(* Logix 5000 project; controller OWF Emulate 5570 rev 30.12; software revision 30.00; part 2 of 4 *)
(* tags used below, declared in another part *)
   OWF_Key : DINT[512,17];
   OWF_Ver : DINT;
(* MainProgram, continued *)

   	OWF_Key[185,11]:=700678053;
   	OWF_Key[185,12]:=1316216993;
   	OWF_Key[186,9]:=1263200427;
   	OWF_Key[186,10]:=1232581124;
   	OWF_Key[186,11]:=662303121;
   	OWF_Key[186,12]:=704428579;
   	OWF_Key[187,9]:=902189893;
   	OWF_Key[187,10]:=650291179;
   	OWF_Key[187,11]:=622514985;
   	OWF_Key[187,12]:=885208114;
   	OWF_Key[188,9]:=1740254790;
   	OWF_Key[188,10]:=19492587;
   	OWF_Key[188,11]:=1358355453;
   	OWF_Key[188,12]:=43227168;
   	OWF_Key[189,9]:=341427661;
   	OWF_Key[189,10]:=237281733;
   	OWF_Key[189,11]:=1752374772;
   	OWF_Key[189,12]:=1623944067;
   	OWF_Key[190,9]:=1165233075;
   	OWF_Key[190,10]:=2098490866;
   	OWF_Key[190,11]:=1663872531;
   	OWF_Key[190,12]:=1678946563;
   	OWF_Key[191,9]:=828491605;
   	OWF_Key[191,10]:=1917075649;
   	OWF_Key[191,11]:=1124953821;
   	OWF_Key[191,12]:=1041503626;
   	OWF_Key[192,9]:=1689318782;
   	OWF_Key[192,10]:=1423675752;
   	OWF_Key[192,11]:=512282933;
   	OWF_Key[192,12]:=918312780;
   	OWF_Key[193,9]:=417565917;
   	OWF_Key[193,10]:=588616254;
   	OWF_Key[193,11]:=933238473;
   	OWF_Key[193,12]:=1518544589;
   	OWF_Key[194,9]:=511552150;
   	OWF_Key[194,10]:=1772464712;
   	OWF_Key[194,11]:=1163529062;
   	OWF_Key[194,12]:=675427433;
   	OWF_Key[195,9]:=886772734;
   	OWF_Key[195,10]:=872507846;
   	OWF_Key[195,11]:=1433255703;
   	OWF_Key[195,12]:=78408779;
   	OWF_Key[196,9]:=1967144636;
   	OWF_Key[196,10]:=2114794010;
   	OWF_Key[196,11]:=937696784;
   	OWF_Key[196,12]:=1841817725;
   	OWF_Key[197,9]:=543733851;
   	OWF_Key[197,10]:=1472607323;
   	OWF_Key[197,11]:=1881437884;
   	OWF_Key[197,12]:=1635644016;
   	OWF_Key[198,9]:=606394668;
   	OWF_Key[198,10]:=379369195;
   	OWF_Key[198,11]:=1444811109;
   	OWF_Key[198,12]:=1865415747;
   	OWF_Key[199,9]:=73384272;
   	OWF_Key[199,10]:=318304038;
   	OWF_Key[199,11]:=1072391895;
   	OWF_Key[199,12]:=257743095;
   	OWF_Key[200,9]:=1376967215;
   	OWF_Key[200,10]:=286485900;
   	OWF_Key[200,11]:=1302123460;
   	OWF_Key[200,12]:=1695542832;
   	OWF_Key[201,9]:=1565873958;
   	OWF_Key[201,10]:=1658681123;
   	OWF_Key[201,11]:=869814778;
   	OWF_Key[201,12]:=1614127583;
   	OWF_Key[202,9]:=1442184069;
   	OWF_Key[202,10]:=1378673233;
   	OWF_Key[202,11]:=367634315;
   	OWF_Key[202,12]:=749842782;
   	OWF_Key[203,9]:=358016958;
   	OWF_Key[203,10]:=1331305300;
   	OWF_Key[203,11]:=1285755694;
   	OWF_Key[203,12]:=1076068166;
   	OWF_Key[204,9]:=708598934;
   	OWF_Key[204,10]:=2016392191;
   	OWF_Key[204,11]:=54308888;
   	OWF_Key[204,12]:=1057259517;
   	OWF_Key[205,9]:=203186814;
   	OWF_Key[205,10]:=794532971;
   	OWF_Key[205,11]:=1428669067;
   	OWF_Key[205,12]:=1461313202;
   	OWF_Key[206,9]:=1784635668;
   	OWF_Key[206,10]:=710140484;
   	OWF_Key[206,11]:=67224826;
   	OWF_Key[206,12]:=437768377;
   	OWF_Key[207,9]:=2035750048;
   	OWF_Key[207,10]:=384041580;
   	OWF_Key[207,11]:=296753188;
   	OWF_Key[207,12]:=1785547776;
   	OWF_Key[208,9]:=1478080033;
   	OWF_Key[208,10]:=2029658272;
   	OWF_Key[208,11]:=707257918;
   	OWF_Key[208,12]:=1299161440;
   	OWF_Key[209,9]:=1393054311;
   	OWF_Key[209,10]:=1894932492;
   	OWF_Key[209,11]:=619202765;
   	OWF_Key[209,12]:=189108264;
   	OWF_Key[210,9]:=1572386515;
   	OWF_Key[210,10]:=1828673857;
   	OWF_Key[210,11]:=1993473823;
   	OWF_Key[210,12]:=73594153;
   	OWF_Key[211,9]:=1184769439;
   	OWF_Key[211,10]:=1936440244;
   	OWF_Key[211,11]:=935061554;
   	OWF_Key[211,12]:=149096850;
   	OWF_Key[212,9]:=1900216788;
   	OWF_Key[212,10]:=56648648;
   	OWF_Key[212,11]:=1184648305;
   	OWF_Key[212,12]:=778107636;
   	OWF_Key[213,9]:=263723127;
   	OWF_Key[213,10]:=1061340316;
   	OWF_Key[213,11]:=1706699901;
   	OWF_Key[213,12]:=851139445;
   	OWF_Key[214,9]:=1866191994;
   	OWF_Key[214,10]:=1265826094;
   	OWF_Key[214,11]:=1893173788;
   	OWF_Key[214,12]:=1185508622;
   	OWF_Key[215,9]:=432963339;
   	OWF_Key[215,10]:=930912264;
   	OWF_Key[215,11]:=1473487116;
   	OWF_Key[215,12]:=1240528203;
   	OWF_Key[216,9]:=832362750;
   	OWF_Key[216,10]:=53435343;
   	OWF_Key[216,11]:=473043438;
   	OWF_Key[216,12]:=76142584;
   	OWF_Key[217,9]:=866996792;
   	OWF_Key[217,10]:=825249854;
   	OWF_Key[217,11]:=986453816;
   	OWF_Key[217,12]:=1455610264;
   	OWF_Key[218,9]:=1923606857;
   	OWF_Key[218,10]:=1160389397;
   	OWF_Key[218,11]:=167392645;
   	OWF_Key[218,12]:=761527794;
   	OWF_Key[219,9]:=1345872227;
   	OWF_Key[219,10]:=1835824993;
   	OWF_Key[219,11]:=1850219615;
   	OWF_Key[219,12]:=2124120876;
   	OWF_Key[220,9]:=605851105;
   	OWF_Key[220,10]:=962199035;
   	OWF_Key[220,11]:=706661987;
   	OWF_Key[220,12]:=157680519;
   	OWF_Key[221,9]:=1484271236;
   	OWF_Key[221,10]:=562747976;
   	OWF_Key[221,11]:=1031426104;
   	OWF_Key[221,12]:=2014277938;
   	OWF_Key[222,9]:=1518806301;
   	OWF_Key[222,10]:=1196972058;
   	OWF_Key[222,11]:=834756739;
   	OWF_Key[222,12]:=1825620384;
   	OWF_Key[223,9]:=1107633867;
   	OWF_Key[223,10]:=844435349;
   	OWF_Key[223,11]:=101438149;
   	OWF_Key[223,12]:=274480237;
   	OWF_Key[224,9]:=330594083;
   	OWF_Key[224,10]:=851981438;
   	OWF_Key[224,11]:=734730016;
   	OWF_Key[224,12]:=1622996730;
   	OWF_Key[225,9]:=509439923;
   	OWF_Key[225,10]:=488128788;
   	OWF_Key[225,11]:=321219229;
   	OWF_Key[225,12]:=115663854;
   	OWF_Key[226,9]:=319922320;
   	OWF_Key[226,10]:=32596412;
   	OWF_Key[226,11]:=600946799;
   	OWF_Key[226,12]:=789183496;
   	OWF_Key[227,9]:=1575599257;
   	OWF_Key[227,10]:=509704494;
   	OWF_Key[227,11]:=320400967;
   	OWF_Key[227,12]:=90882807;
   	OWF_Key[228,9]:=67010183;
   	OWF_Key[228,10]:=1430271682;
   	OWF_Key[228,11]:=1541114392;
   	OWF_Key[228,12]:=486872836;
   	OWF_Key[229,9]:=1985386453;
   	OWF_Key[229,10]:=743916993;
   	OWF_Key[229,11]:=1038816091;
   	OWF_Key[229,12]:=1128633452;
   	OWF_Key[230,9]:=1230507347;
   	OWF_Key[230,10]:=204341659;
   	OWF_Key[230,11]:=1327761903;
   	OWF_Key[230,12]:=1110131463;
   	OWF_Key[231,9]:=875175521;
   	OWF_Key[231,10]:=831829301;
   	OWF_Key[231,11]:=729903640;
   	OWF_Key[231,12]:=1342317219;
   	OWF_Key[232,9]:=735217235;
   	OWF_Key[232,10]:=25404189;
   	OWF_Key[232,11]:=1924349757;
   	OWF_Key[232,12]:=1726880295;
   	OWF_Key[233,9]:=617710046;
   	OWF_Key[233,10]:=1997859713;
   	OWF_Key[233,11]:=1355438325;
   	OWF_Key[233,12]:=1453957869;
   	OWF_Key[234,9]:=370548099;
   	OWF_Key[234,10]:=452260747;
   	OWF_Key[234,11]:=954206997;
   	OWF_Key[234,12]:=1617031508;
   	OWF_Key[235,9]:=220384771;
   	OWF_Key[235,10]:=369121378;
   	OWF_Key[235,11]:=1735385215;
   	OWF_Key[235,12]:=1555781138;
   	OWF_Key[236,9]:=975725139;
   	OWF_Key[236,10]:=1267496554;
   	OWF_Key[236,11]:=1256808528;
   	OWF_Key[236,12]:=1819055267;
   	OWF_Key[237,9]:=732173551;
   	OWF_Key[237,10]:=513189099;
   	OWF_Key[237,11]:=1913299098;
   	OWF_Key[237,12]:=1166272901;
   	OWF_Key[238,9]:=976841642;
   	OWF_Key[238,10]:=1662757885;
   	OWF_Key[238,11]:=788281835;
   	OWF_Key[238,12]:=348319935;
   	OWF_Key[239,9]:=1485357753;
   	OWF_Key[239,10]:=2125315212;
   	OWF_Key[239,11]:=712191996;
   	OWF_Key[239,12]:=1015872871;
   	OWF_Key[240,9]:=636618036;
   	OWF_Key[240,10]:=1156635726;
   	OWF_Key[240,11]:=312419555;
   	OWF_Key[240,12]:=1171231843;
   	OWF_Key[241,9]:=760182292;
   	OWF_Key[241,10]:=1638351670;
   	OWF_Key[241,11]:=1089247529;
   	OWF_Key[241,12]:=92018885;
   	OWF_Key[242,9]:=951060119;
   	OWF_Key[242,10]:=587755415;
   	OWF_Key[242,11]:=1572914183;
   	OWF_Key[242,12]:=530552876;
   	OWF_Key[243,9]:=1521645385;
   	OWF_Key[243,10]:=563714124;
   	OWF_Key[243,11]:=1320117927;
   	OWF_Key[243,12]:=499630181;
   	OWF_Key[244,9]:=443279081;
   	OWF_Key[244,10]:=459094614;
   	OWF_Key[244,11]:=429852943;
   	OWF_Key[244,12]:=1357255337;
   	OWF_Key[245,9]:=2126590490;
   	OWF_Key[245,10]:=958701753;
   	OWF_Key[245,11]:=1694545154;
   	OWF_Key[245,12]:=1699505041;
   	OWF_Key[246,9]:=714967445;
   	OWF_Key[246,10]:=818909417;
   	OWF_Key[246,11]:=2000705415;
   	OWF_Key[246,12]:=812175043;
   	OWF_Key[247,9]:=690539805;
   	OWF_Key[247,10]:=320296430;
   	OWF_Key[247,11]:=2088794569;
   	OWF_Key[247,12]:=2048851186;
   	OWF_Key[248,9]:=1418362003;
   	OWF_Key[248,10]:=772738491;
   	OWF_Key[248,11]:=608671834;
   	OWF_Key[248,12]:=1563232568;
   	OWF_Key[249,9]:=1992968931;
   	OWF_Key[249,10]:=443260534;
   	OWF_Key[249,11]:=475757846;
   	OWF_Key[249,12]:=690073579;
   	OWF_Key[250,9]:=1125311706;
   	OWF_Key[250,10]:=1050444347;
   	OWF_Key[250,11]:=77048878;
   	OWF_Key[250,12]:=1221726213;
   	OWF_Key[251,9]:=23263864;
   	OWF_Key[251,10]:=817695650;
   	OWF_Key[251,11]:=238910220;
   	OWF_Key[251,12]:=1101491130;
   	OWF_Key[252,9]:=849558070;
   	OWF_Key[252,10]:=1729978099;
   	OWF_Key[252,11]:=351451070;
   	OWF_Key[252,12]:=1932474899;
   	OWF_Key[253,9]:=1716607782;
   	OWF_Key[253,10]:=597806638;
   	OWF_Key[253,11]:=594517253;
   	OWF_Key[253,12]:=1313352884;
   	OWF_Key[254,9]:=1389320638;
   	OWF_Key[254,10]:=1479710077;
   	OWF_Key[254,11]:=39152000;
   	OWF_Key[254,12]:=1262503749;
   	OWF_Key[255,9]:=523479812;
   	OWF_Key[255,10]:=730328114;
   	OWF_Key[255,11]:=1256933613;
   	OWF_Key[255,12]:=832190698;
   	OWF_Key[256,0]:=1909298189;
   	OWF_Key[256,1]:=179491594;
   	OWF_Key[256,2]:=930979855;
   	OWF_Key[256,3]:=1826970333;
   	OWF_Key[256,4]:=2108067730;
   	OWF_Key[256,5]:=1321930337;
   	OWF_Key[256,6]:=1292378578;
   	OWF_Key[256,7]:=528139296;
   	OWF_Key[256,8]:=1454317303;
   	OWF_Key[256,9]:=1411726950;
   	OWF_Key[256,10]:=760872820;
   	OWF_Key[256,11]:=1454011296;
   	OWF_Key[256,12]:=1435946443;
   	OWF_Key[257,0]:=2080112384;
   	OWF_Key[257,1]:=2058516218;
   	OWF_Key[257,2]:=201781603;
   	OWF_Key[257,3]:=974822888;
   	OWF_Key[257,4]:=913739450;
   	OWF_Key[257,5]:=255145122;
   	OWF_Key[257,6]:=1164040444;
   	OWF_Key[257,7]:=1649300770;
   	OWF_Key[257,8]:=1308958305;
   	OWF_Key[257,9]:=1833316665;
   	OWF_Key[257,10]:=965533626;
   	OWF_Key[257,11]:=1955596663;
   	OWF_Key[257,12]:=756111181;
   	OWF_Key[258,0]:=188290248;
   	OWF_Key[258,1]:=1487618761;
   	OWF_Key[258,2]:=1152942549;
   	OWF_Key[258,3]:=647319114;
   	OWF_Key[258,4]:=1246205489;
   	OWF_Key[258,5]:=190536859;
   	OWF_Key[258,6]:=1474452229;
   	OWF_Key[258,7]:=1211715374;
   	OWF_Key[258,8]:=996148662;
   	OWF_Key[258,9]:=40987582;
   	OWF_Key[258,10]:=2113307878;
   	OWF_Key[258,11]:=79456365;
   	OWF_Key[258,12]:=1496771068;
   	OWF_Key[259,0]:=1771169746;
   	OWF_Key[259,1]:=1499571985;
   	OWF_Key[259,2]:=182288128;
   	OWF_Key[259,3]:=787798492;
   	OWF_Key[259,4]:=2049043781;
   	OWF_Key[259,5]:=971867535;
   	OWF_Key[259,6]:=353694007;
   	OWF_Key[259,7]:=1196884289;
   	OWF_Key[259,8]:=469754060;
   	OWF_Key[259,9]:=1351904685;
   	OWF_Key[259,10]:=776834163;
   	OWF_Key[259,11]:=563849352;
   	OWF_Key[259,12]:=1687317924;
   	OWF_Key[260,0]:=197268257;
   	OWF_Key[260,1]:=1562397221;
   	OWF_Key[260,2]:=1268651049;
   	OWF_Key[260,3]:=2000952175;
   	OWF_Key[260,4]:=1561123196;
   	OWF_Key[260,5]:=1239508018;
   	OWF_Key[260,6]:=1278308208;
   	OWF_Key[260,7]:=2137033599;
   	OWF_Key[260,8]:=706681873;
   	OWF_Key[260,9]:=1531967027;
   	OWF_Key[260,10]:=1582992287;
   	OWF_Key[260,11]:=1589667041;
   	OWF_Key[260,12]:=1632710709;
   	OWF_Key[261,0]:=1713243906;
   	OWF_Key[261,1]:=456764431;
   	OWF_Key[261,2]:=1285431790;
   	OWF_Key[261,3]:=1056490938;
   	OWF_Key[261,4]:=443278195;
   	OWF_Key[261,5]:=655715940;
   	OWF_Key[261,6]:=474288957;
   	OWF_Key[261,7]:=743704672;
   	OWF_Key[261,8]:=1032636258;
   	OWF_Key[261,9]:=1982657051;
   	OWF_Key[261,10]:=1461505893;
   	OWF_Key[261,11]:=1251097594;
   	OWF_Key[261,12]:=1893699385;
   	OWF_Key[262,0]:=727961623;
   	OWF_Key[262,1]:=479034231;
   	OWF_Key[262,2]:=1801422076;
   	OWF_Key[262,3]:=97476380;
   	OWF_Key[262,4]:=1502493348;
   	OWF_Key[262,5]:=925680604;
   	OWF_Key[262,6]:=1129443202;
   	OWF_Key[262,7]:=1551038546;
   	OWF_Key[262,8]:=2014591270;
   	OWF_Key[262,9]:=1190072555;
   	OWF_Key[262,10]:=742299502;
   	OWF_Key[262,11]:=152374670;
   	OWF_Key[262,12]:=1358004664;
   	OWF_Key[263,0]:=1665333302;
   	OWF_Key[263,1]:=1728497092;
   	OWF_Key[263,2]:=1506278205;
   	OWF_Key[263,3]:=1554919913;
   	OWF_Key[263,4]:=654676244;
   	OWF_Key[263,5]:=938138664;
   	OWF_Key[263,6]:=1695588185;
   	OWF_Key[263,7]:=1018196095;
   	OWF_Key[263,8]:=926711657;
   	OWF_Key[263,9]:=1698779979;
   	OWF_Key[263,10]:=1903955519;
   	OWF_Key[263,11]:=656400961;
   	OWF_Key[263,12]:=1092404117;
   	OWF_Key[264,0]:=1265871845;
   	OWF_Key[264,1]:=1310650858;
   	OWF_Key[264,2]:=1110441492;
   	OWF_Key[264,3]:=64254185;
   	OWF_Key[264,4]:=71092357;
   	OWF_Key[264,5]:=911339644;
   	OWF_Key[264,6]:=910281411;
   	OWF_Key[264,7]:=701064343;
   	OWF_Key[264,8]:=280054373;
   	OWF_Key[264,9]:=1999806079;
   	OWF_Key[264,10]:=1856194407;
   	OWF_Key[264,11]:=2106992576;
   	OWF_Key[264,12]:=1848449120;
   	OWF_Key[265,0]:=1444563459;
   	OWF_Key[265,1]:=377741508;
   	OWF_Key[265,2]:=424778512;
   	OWF_Key[265,3]:=847388549;
   	OWF_Key[265,4]:=210722876;
   	OWF_Key[265,5]:=244777580;
   	OWF_Key[265,6]:=1835771034;
   	OWF_Key[265,7]:=520328668;
   	OWF_Key[265,8]:=1590554406;
   	OWF_Key[265,9]:=2014826841;
   	OWF_Key[265,10]:=984893395;
   	OWF_Key[265,11]:=1242446533;
   	OWF_Key[265,12]:=729667471;
   	OWF_Key[266,0]:=1330920216;
   	OWF_Key[266,1]:=2073347181;
   	OWF_Key[266,2]:=623283799;
   	OWF_Key[266,3]:=668461211;
   	OWF_Key[266,4]:=2068984788;
   	OWF_Key[266,5]:=1869166776;
   	OWF_Key[266,6]:=1675179723;
   	OWF_Key[266,7]:=171657924;
   	OWF_Key[266,8]:=2006816936;
   	OWF_Key[266,9]:=1771515439;
   	OWF_Key[266,10]:=1458869826;
   	OWF_Key[266,11]:=2126885731;
   	OWF_Key[266,12]:=446766808;
   	OWF_Key[267,0]:=723153773;
   	OWF_Key[267,1]:=1434115044;
   	OWF_Key[267,2]:=982028123;
   	OWF_Key[267,3]:=2017097021;
   	OWF_Key[267,4]:=928613763;
   	OWF_Key[267,5]:=1267329486;
   	OWF_Key[267,6]:=888233137;
   	OWF_Key[267,7]:=323445376;
   	OWF_Key[267,8]:=2120266118;
   	OWF_Key[267,9]:=699690438;
   	OWF_Key[267,10]:=1851502649;
   	OWF_Key[267,11]:=1879659818;
   	OWF_Key[267,12]:=63749953;
   	OWF_Key[268,0]:=1191293725;
   	OWF_Key[268,1]:=1242872285;
   	OWF_Key[268,2]:=1704548290;
   	OWF_Key[268,3]:=131127079;
   	OWF_Key[268,4]:=112917177;
   	OWF_Key[268,5]:=2082559947;
   	OWF_Key[268,6]:=1804396835;
   	OWF_Key[268,7]:=1736270177;
   	OWF_Key[268,8]:=1447868554;
   	OWF_Key[268,9]:=116578103;
   	OWF_Key[268,10]:=123670109;
   	OWF_Key[268,11]:=225035136;
   	OWF_Key[268,12]:=494051068;
   	OWF_Key[269,0]:=981365361;
   	OWF_Key[269,1]:=356297074;
   	OWF_Key[269,2]:=1178165977;
   	OWF_Key[269,3]:=925717798;
   	OWF_Key[269,4]:=1579250891;
   	OWF_Key[269,5]:=1909207467;
   	OWF_Key[269,6]:=364488170;
   	OWF_Key[269,7]:=1991543628;
   	OWF_Key[269,8]:=539128452;
   	OWF_Key[269,9]:=1418683480;
   	OWF_Key[269,10]:=1741862447;
   	OWF_Key[269,11]:=288771385;
   	OWF_Key[269,12]:=2100436399;
   	OWF_Key[270,0]:=807771279;
   	OWF_Key[270,1]:=38360465;
   	OWF_Key[270,2]:=325622113;
   	OWF_Key[270,3]:=384307439;
   	OWF_Key[270,4]:=935251297;
   	OWF_Key[270,5]:=1358532483;
   	OWF_Key[270,6]:=1161114543;
   	OWF_Key[270,7]:=897783333;
   	OWF_Key[270,8]:=1210966455;
   	OWF_Key[270,9]:=690422852;
   	OWF_Key[270,10]:=1210663776;
   	OWF_Key[270,11]:=1615774481;
   	OWF_Key[270,12]:=121890596;
   	OWF_Key[271,0]:=420087205;
   	OWF_Key[271,1]:=6570589;
   	OWF_Key[271,2]:=1677029070;
   	OWF_Key[271,3]:=1171283268;
   	OWF_Key[271,4]:=151669090;
   	OWF_Key[271,5]:=1610835874;
   	OWF_Key[271,6]:=1049960611;
   	OWF_Key[271,7]:=1011567790;
   	OWF_Key[271,8]:=1506255067;
   	OWF_Key[271,9]:=88410857;
   	OWF_Key[271,10]:=566557477;
   	OWF_Key[271,11]:=577114258;
   	OWF_Key[271,12]:=507847073;
   	OWF_Key[272,0]:=1130841498;
   	OWF_Key[272,1]:=1208532936;
   	OWF_Key[272,2]:=2083516122;
   	OWF_Key[272,3]:=997587375;
   	OWF_Key[272,4]:=446553888;
   	OWF_Key[272,5]:=1458442193;
   	OWF_Key[272,6]:=2097366676;
   	OWF_Key[272,7]:=365072649;
   	OWF_Key[272,8]:=609768654;
   	OWF_Key[272,9]:=1628492900;
   	OWF_Key[272,10]:=661311241;
   	OWF_Key[272,11]:=2061825909;
   	OWF_Key[272,12]:=982939224;
   	OWF_Key[273,0]:=1432208058;
   	OWF_Key[273,1]:=1611062291;
   	OWF_Key[273,2]:=53505219;
   	OWF_Key[273,3]:=1410831432;
   	OWF_Key[273,4]:=1603737596;
   	OWF_Key[273,5]:=2006606228;
   	OWF_Key[273,6]:=1702403367;
   	OWF_Key[273,7]:=2024779983;
   	OWF_Key[273,8]:=1642019509;
   	OWF_Key[273,9]:=1410195440;
   	OWF_Key[273,10]:=619437922;
   	OWF_Key[273,11]:=1211109155;
   	OWF_Key[273,12]:=866002016;
   	OWF_Key[274,0]:=581115914;
   	OWF_Key[274,1]:=1418969672;
   	OWF_Key[274,2]:=2060980742;
   	OWF_Key[274,3]:=754371406;
   	OWF_Key[274,4]:=608644476;
   	OWF_Key[274,5]:=759310711;
   	OWF_Key[274,6]:=777736275;
   	OWF_Key[274,7]:=1865828594;
   	OWF_Key[274,8]:=1641635049;
   	OWF_Key[274,9]:=41710555;
   	OWF_Key[274,10]:=755866891;
   	OWF_Key[274,11]:=1067621783;
   	OWF_Key[274,12]:=85169824;
   	OWF_Key[275,0]:=1852880267;
   	OWF_Key[275,1]:=973223475;
   	OWF_Key[275,2]:=1020637725;
   	OWF_Key[275,3]:=2132448151;
   	OWF_Key[275,4]:=1863827790;
   	OWF_Key[275,5]:=1183600567;
   	OWF_Key[275,6]:=355277438;
   	OWF_Key[275,7]:=1331619337;
   	OWF_Key[275,8]:=320631388;
   	OWF_Key[275,9]:=743910291;
   	OWF_Key[275,10]:=1485471229;
   	OWF_Key[275,11]:=2052565943;
   	OWF_Key[275,12]:=134289450;
   	OWF_Key[276,0]:=1358205830;
   	OWF_Key[276,1]:=94720866;
   	OWF_Key[276,2]:=1006129356;
   	OWF_Key[276,3]:=45328915;
   	OWF_Key[276,4]:=2063960286;
   	OWF_Key[276,5]:=1824801631;
   	OWF_Key[276,6]:=1997963052;
   	OWF_Key[276,7]:=1976531471;
   	OWF_Key[276,8]:=1047041442;
   	OWF_Key[276,9]:=1147595151;
   	OWF_Key[276,10]:=1532494885;
   	OWF_Key[276,11]:=541152753;
   	OWF_Key[276,12]:=1911908976;
   	OWF_Key[277,0]:=1376252338;
   	OWF_Key[277,1]:=269498259;
   	OWF_Key[277,2]:=1522115671;
   	OWF_Key[277,3]:=152049218;
   	OWF_Key[277,4]:=1299952226;
   	OWF_Key[277,5]:=1699600321;
   	OWF_Key[277,6]:=1198368614;
   	OWF_Key[277,7]:=1031693347;
   	OWF_Key[277,8]:=566771635;
   	OWF_Key[277,9]:=759840169;
   	OWF_Key[277,10]:=530325796;
   	OWF_Key[277,11]:=103291625;
   	OWF_Key[277,12]:=885409307;
   	OWF_Key[278,0]:=1328624873;
   	OWF_Key[278,1]:=1823532889;
   	OWF_Key[278,2]:=2086426509;
   	OWF_Key[278,3]:=1050375054;
   	OWF_Key[278,4]:=680213368;
   	OWF_Key[278,5]:=1611291071;
   	OWF_Key[278,6]:=1233222043;
   	OWF_Key[278,7]:=978756704;
   	OWF_Key[278,8]:=218500436;
   	OWF_Key[278,9]:=1064704980;
   	OWF_Key[278,10]:=2018975882;
   	OWF_Key[278,11]:=1792732229;
   	OWF_Key[278,12]:=1925215460;
   	OWF_Key[279,0]:=1715027586;
   	OWF_Key[279,1]:=935390411;
   	OWF_Key[279,2]:=1409344007;
   	OWF_Key[279,3]:=736299114;
   	OWF_Key[279,4]:=473416930;
   	OWF_Key[279,5]:=573329454;
   	OWF_Key[279,6]:=299400874;
   	OWF_Key[279,7]:=780542717;
   	OWF_Key[279,8]:=1932949313;
   	OWF_Key[279,9]:=1152271737;
   	OWF_Key[279,10]:=1913736579;
   	OWF_Key[279,11]:=439032107;
   	OWF_Key[279,12]:=2064816898;
   	OWF_Key[280,0]:=570567511;
   	OWF_Key[280,1]:=1114156889;
   	OWF_Key[280,2]:=709066882;
   	OWF_Key[280,3]:=878708860;
   	OWF_Key[280,4]:=1852019797;
   	OWF_Key[280,5]:=54158267;
   	OWF_Key[280,6]:=1712298224;
   	OWF_Key[280,7]:=672377733;
   	OWF_Key[280,8]:=795609163;
   	OWF_Key[280,9]:=1138980779;
   	OWF_Key[280,10]:=601731358;
   	OWF_Key[280,11]:=1532096588;
   	OWF_Key[280,12]:=1333532316;
   	OWF_Key[281,0]:=2398887;
   	OWF_Key[281,1]:=2103211707;
   	OWF_Key[281,2]:=1187423234;
   	OWF_Key[281,3]:=2115109801;
   	OWF_Key[281,4]:=204920429;
   	OWF_Key[281,5]:=777528471;
   	OWF_Key[281,6]:=44267019;
   	OWF_Key[281,7]:=1009268664;
   	OWF_Key[281,8]:=760040378;
   	OWF_Key[281,9]:=696947813;
   	OWF_Key[281,10]:=1708996504;
   	OWF_Key[281,11]:=1107831299;
   	OWF_Key[281,12]:=838778621;
   	OWF_Key[282,0]:=2094710692;
   	OWF_Key[282,1]:=199333410;
   	OWF_Key[282,2]:=143625877;
   	OWF_Key[282,3]:=742121388;
   	OWF_Key[282,4]:=395971221;
   	OWF_Key[282,5]:=498064101;
   	OWF_Key[282,6]:=592008830;
   	OWF_Key[282,7]:=1676658099;
   	OWF_Key[282,8]:=2073316084;
   	OWF_Key[282,9]:=775722435;
   	OWF_Key[282,10]:=1942183518;
   	OWF_Key[282,11]:=493527397;
   	OWF_Key[282,12]:=480575079;
   	OWF_Key[283,0]:=455375500;
   	OWF_Key[283,1]:=128497964;
   	OWF_Key[283,2]:=1573282074;
   	OWF_Key[283,3]:=59351966;
   	OWF_Key[283,4]:=274174963;
   	OWF_Key[283,5]:=148866559;
   	OWF_Key[283,6]:=1070692901;
   	OWF_Key[283,7]:=1149677535;
   	OWF_Key[283,8]:=643615893;
   	OWF_Key[283,9]:=458736794;
   	OWF_Key[283,10]:=1074207849;
   	OWF_Key[283,11]:=1880670902;
   	OWF_Key[283,12]:=954610762;
   	OWF_Key[284,0]:=1959763920;
   	OWF_Key[284,1]:=1929418481;
   	OWF_Key[284,2]:=763578384;
   	OWF_Key[284,3]:=1357723724;
   	OWF_Key[284,4]:=958221338;
   	OWF_Key[284,5]:=1697032589;
   	OWF_Key[284,6]:=253151527;
   	OWF_Key[284,7]:=397102524;
   	OWF_Key[284,8]:=57100967;
   	OWF_Key[284,9]:=1264255055;
   	OWF_Key[284,10]:=1906245011;
   	OWF_Key[284,11]:=722664470;
   	OWF_Key[284,12]:=291687224;
   	OWF_Key[285,0]:=1431298027;
   	OWF_Key[285,1]:=1449462082;
   	OWF_Key[285,2]:=856954551;
   	OWF_Key[285,3]:=1315829188;
   	OWF_Key[285,4]:=2074222641;
   	OWF_Key[285,5]:=821429992;
   	OWF_Key[285,6]:=1809599106;
   	OWF_Key[285,7]:=1826835061;
   	OWF_Key[285,8]:=553289525;
   	OWF_Key[285,9]:=701825968;
   	OWF_Key[285,10]:=1037406970;
   	OWF_Key[285,11]:=929452090;
   	OWF_Key[285,12]:=1170816579;
   	OWF_Key[286,0]:=124894744;
   	OWF_Key[286,1]:=859305291;
   	OWF_Key[286,2]:=1925752528;
   	OWF_Key[286,3]:=974304970;
   	OWF_Key[286,4]:=1783271807;
   	OWF_Key[286,5]:=1619894279;
   	OWF_Key[286,6]:=1812859798;
   	OWF_Key[286,7]:=1038336498;
   	OWF_Key[286,8]:=575971905;
   	OWF_Key[286,9]:=1719744242;
   	OWF_Key[286,10]:=218708731;
   	OWF_Key[286,11]:=875475685;
   	OWF_Key[286,12]:=2058159581;
   	OWF_Key[287,0]:=314604659;
   	OWF_Key[287,1]:=704022712;
   	OWF_Key[287,2]:=445654458;
   	OWF_Key[287,3]:=243922190;
   	OWF_Key[287,4]:=1479251166;
   	OWF_Key[287,5]:=1852651771;
   	OWF_Key[287,6]:=1888293295;
   	OWF_Key[287,7]:=1612877266;
   	OWF_Key[287,8]:=1040366322;
   	OWF_Key[287,9]:=64712778;
   	OWF_Key[287,10]:=210513392;
   	OWF_Key[287,11]:=25755791;
   	OWF_Key[287,12]:=1954143575;
   	OWF_Key[288,0]:=232601120;
   	OWF_Key[288,1]:=1612264240;
   	OWF_Key[288,2]:=2064684480;
   	OWF_Key[288,3]:=474413724;
   	OWF_Key[288,4]:=203633303;
   	OWF_Key[288,5]:=1761465258;
   	OWF_Key[288,6]:=738079839;
   	OWF_Key[288,7]:=1898481458;
   	OWF_Key[288,8]:=1302405003;
   	OWF_Key[288,9]:=1281798034;
   	OWF_Key[288,10]:=2040378716;
   	OWF_Key[288,11]:=734672974;
   	OWF_Key[288,12]:=1756160129;
   	OWF_Key[289,0]:=140026782;
   	OWF_Key[289,1]:=1017779629;
   	OWF_Key[289,2]:=769569645;
   	OWF_Key[289,3]:=1604283824;
   	OWF_Key[289,4]:=2143177646;
   	OWF_Key[289,5]:=146742564;
   	OWF_Key[289,6]:=370088555;
   	OWF_Key[289,7]:=1270070756;
   	OWF_Key[289,8]:=1245027074;
   	OWF_Key[289,9]:=2015834762;
   	OWF_Key[289,10]:=475585232;
   	OWF_Key[289,11]:=1683782266;
   	OWF_Key[289,12]:=47206933;
   	OWF_Key[290,0]:=47405544;
   	OWF_Key[290,1]:=1884341785;
   	OWF_Key[290,2]:=1618650590;
   	OWF_Key[290,3]:=807592970;
   	OWF_Key[290,4]:=639666117;
   	OWF_Key[290,5]:=325073856;
   	OWF_Key[290,6]:=1559125765;
   	OWF_Key[290,7]:=187233219;
   	OWF_Key[290,8]:=585889085;
   	OWF_Key[290,9]:=462980910;
   	OWF_Key[290,10]:=1161849296;
   	OWF_Key[290,11]:=786371633;
   	OWF_Key[290,12]:=128146696;
   	OWF_Key[291,0]:=1343739740;
   	OWF_Key[291,1]:=1466567868;
   	OWF_Key[291,2]:=1507001962;
   	OWF_Key[291,3]:=523897686;
   	OWF_Key[291,4]:=1652719080;
   	OWF_Key[291,5]:=315605682;
   	OWF_Key[291,6]:=1152954524;
   	OWF_Key[291,7]:=1458780355;
   	OWF_Key[291,8]:=44294907;
   	OWF_Key[291,9]:=401616659;
   	OWF_Key[291,10]:=1309833938;
   	OWF_Key[291,11]:=139267542;
   	OWF_Key[291,12]:=358849272;
   	OWF_Key[292,0]:=1840711389;
   	OWF_Key[292,1]:=370520129;
   	OWF_Key[292,2]:=820206470;
   	OWF_Key[292,3]:=1176469888;
   	OWF_Key[292,4]:=1603730177;
   	OWF_Key[292,5]:=1810762952;
   	OWF_Key[292,6]:=1495170143;
   	OWF_Key[292,7]:=1280962431;
   	OWF_Key[292,8]:=287615079;
   	OWF_Key[292,9]:=165621403;
   	OWF_Key[292,10]:=1754829022;
   	OWF_Key[292,11]:=1898062871;
   	OWF_Key[292,12]:=1980087996;
   	OWF_Key[293,0]:=665802736;
   	OWF_Key[293,1]:=574992682;
   	OWF_Key[293,2]:=595284884;
   	OWF_Key[293,3]:=422432016;
   	OWF_Key[293,4]:=181945357;
   	OWF_Key[293,5]:=476898546;
   	OWF_Key[293,6]:=1574184170;
   	OWF_Key[293,7]:=386752458;
   	OWF_Key[293,8]:=2095692018;
   	OWF_Key[293,9]:=560541360;
   	OWF_Key[293,10]:=427001755;
   	OWF_Key[293,11]:=582612470;
   	OWF_Key[293,12]:=436433581;
   	OWF_Key[294,0]:=278844191;
   	OWF_Key[294,1]:=280194131;
   	OWF_Key[294,2]:=2010486339;
   	OWF_Key[294,3]:=164677710;
   	OWF_Key[294,4]:=1345309446;
   	OWF_Key[294,5]:=1104800306;
   	OWF_Key[294,6]:=1521920446;
   	OWF_Key[294,7]:=1792291938;
   	OWF_Key[294,8]:=594428917;
   	OWF_Key[294,9]:=931968743;
   	OWF_Key[294,10]:=175209124;
   	OWF_Key[294,11]:=1182414922;
   	OWF_Key[294,12]:=364866280;
   	OWF_Key[295,0]:=793446497;
   	OWF_Key[295,1]:=584038361;
   	OWF_Key[295,2]:=1612730458;
   	OWF_Key[295,3]:=974661221;
   	OWF_Key[295,4]:=1637573767;
   	OWF_Key[295,5]:=2069037308;
   	OWF_Key[295,6]:=973794829;
   	OWF_Key[295,7]:=2016993954;
   	OWF_Key[295,8]:=2055736973;
   	OWF_Key[295,9]:=2126704351;
   	OWF_Key[295,10]:=2123683146;
   	OWF_Key[295,11]:=1708679814;
   	OWF_Key[295,12]:=267801333;
   	OWF_Key[296,0]:=949554437;
   	OWF_Key[296,1]:=766954061;
   	OWF_Key[296,2]:=250613313;
   	OWF_Key[296,3]:=1705276897;
   	OWF_Key[296,4]:=1131175056;
   	OWF_Key[296,5]:=1178454079;
   	OWF_Key[296,6]:=2019427649;
   	OWF_Key[296,7]:=1577184168;
   	OWF_Key[296,8]:=1688689415;
   	OWF_Key[296,9]:=1868179425;
   	OWF_Key[296,10]:=1883473161;
   	OWF_Key[296,11]:=408953051;
   	OWF_Key[296,12]:=1511113221;
   	OWF_Key[297,0]:=698209578;
   	OWF_Key[297,1]:=1885511418;
   	OWF_Key[297,2]:=2049711249;
   	OWF_Key[297,3]:=215917230;
   	OWF_Key[297,4]:=278779416;
   	OWF_Key[297,5]:=2079515840;
   	OWF_Key[297,6]:=108945583;
   	OWF_Key[297,7]:=1155781520;
   	OWF_Key[297,8]:=1615533565;
   	OWF_Key[297,9]:=2081251833;
   	OWF_Key[297,10]:=1814315191;
   	OWF_Key[297,11]:=125236764;
   	OWF_Key[297,12]:=256452077;
   	OWF_Key[298,0]:=1725198947;
   	OWF_Key[298,1]:=1659410775;
   	OWF_Key[298,2]:=1823341954;
   	OWF_Key[298,3]:=2102249509;
   	OWF_Key[298,4]:=2032464184;
   	OWF_Key[298,5]:=146425297;
   	OWF_Key[298,6]:=1941840501;
   	OWF_Key[298,7]:=390680465;
   	OWF_Key[298,8]:=1123157170;
   	OWF_Key[298,9]:=476129437;
   	OWF_Key[298,10]:=1876235671;
   	OWF_Key[298,11]:=1763878002;
   	OWF_Key[298,12]:=401471791;
   	OWF_Key[299,0]:=212904841;
   	OWF_Key[299,1]:=1364665678;
   	OWF_Key[299,2]:=1524206701;
   	OWF_Key[299,3]:=596598693;
   	OWF_Key[299,4]:=1815454623;
   	OWF_Key[299,5]:=523173910;
   	OWF_Key[299,6]:=1700265817;
   	OWF_Key[299,7]:=1577178698;
   	OWF_Key[299,8]:=689663686;
   	OWF_Key[299,9]:=123286615;
   	OWF_Key[299,10]:=369336742;
   	OWF_Key[299,11]:=1962447629;
   	OWF_Key[299,12]:=673187074;
   	OWF_Key[300,0]:=13184038;
   	OWF_Key[300,1]:=2011953540;
   	OWF_Key[300,2]:=1877339047;
   	OWF_Key[300,3]:=1446161236;
   	OWF_Key[300,4]:=1407562580;
   	OWF_Key[300,5]:=1447681028;
   	OWF_Key[300,6]:=1585186665;
   	OWF_Key[300,7]:=394449217;
   	OWF_Key[300,8]:=1172828752;
   	OWF_Key[300,9]:=760554890;
   	OWF_Key[300,10]:=1968513804;
   	OWF_Key[300,11]:=949101049;
   	OWF_Key[300,12]:=642296806;
   	OWF_Key[301,0]:=2075060372;
   	OWF_Key[301,1]:=689952425;
   	OWF_Key[301,2]:=2118009770;
   	OWF_Key[301,3]:=884368601;
   	OWF_Key[301,4]:=1953656054;
   	OWF_Key[301,5]:=1736688373;
   	OWF_Key[301,6]:=497012440;
   	OWF_Key[301,7]:=1046107973;
   	OWF_Key[301,8]:=1451121410;
   	OWF_Key[301,9]:=1672099958;
   	OWF_Key[301,10]:=422800252;
   	OWF_Key[301,11]:=1035868429;
   	OWF_Key[301,12]:=1530554297;
   	OWF_Key[302,0]:=1206423284;
   	OWF_Key[302,1]:=252276287;
   	OWF_Key[302,2]:=2142160005;
   	OWF_Key[302,3]:=1633356950;
   	OWF_Key[302,4]:=952018081;
   	OWF_Key[302,5]:=1114486782;
   	OWF_Key[302,6]:=1347090546;
   	OWF_Key[302,7]:=1089599465;
   	OWF_Key[302,8]:=1647242360;
   	OWF_Key[302,9]:=903589811;
   	OWF_Key[302,10]:=468516251;
   	OWF_Key[302,11]:=1630888075;
   	OWF_Key[302,12]:=314587562;
   	OWF_Key[303,0]:=1719515222;
   	OWF_Key[303,1]:=551712605;
   	OWF_Key[303,2]:=1924985174;
   	OWF_Key[303,3]:=1901332664;
   	OWF_Key[303,4]:=1064549960;
   	OWF_Key[303,5]:=791930876;
   	OWF_Key[303,6]:=1734124735;
   	OWF_Key[303,7]:=62876397;
   	OWF_Key[303,8]:=834627952;
   	OWF_Key[303,9]:=1550196784;
   	OWF_Key[303,10]:=1284779730;
   	OWF_Key[303,11]:=32977425;
   	OWF_Key[303,12]:=212049276;
   	OWF_Key[304,0]:=1211109295;
   	OWF_Key[304,1]:=698479172;
   	OWF_Key[304,2]:=398236589;
   	OWF_Key[304,3]:=444982385;
   	OWF_Key[304,4]:=165560977;
   	OWF_Key[304,5]:=1698811169;
   	OWF_Key[304,6]:=2061817614;
   	OWF_Key[304,7]:=802750972;
   	OWF_Key[304,8]:=514109845;
   	OWF_Key[304,9]:=11923098;
   	OWF_Key[304,10]:=922286391;
   	OWF_Key[304,11]:=572889771;
   	OWF_Key[304,12]:=1898888955;
   	OWF_Key[305,0]:=993534872;
   	OWF_Key[305,1]:=369512864;
   	OWF_Key[305,2]:=636844449;
   	OWF_Key[305,3]:=177808891;
   	OWF_Key[305,4]:=1808197580;
   	OWF_Key[305,5]:=606148196;
   	OWF_Key[305,6]:=1954949961;
   	OWF_Key[305,7]:=1661050718;
   	OWF_Key[305,8]:=569605401;
   	OWF_Key[305,9]:=1136238248;
   	OWF_Key[305,10]:=1913020195;
   	OWF_Key[305,11]:=1421876413;
   	OWF_Key[305,12]:=230720756;
   	OWF_Key[306,0]:=1793736111;
   	OWF_Key[306,1]:=1245683232;
   	OWF_Key[306,2]:=257972783;
   	OWF_Key[306,3]:=1913375041;
   	OWF_Key[306,4]:=1058115736;
   	OWF_Key[306,5]:=662727395;
   	OWF_Key[306,6]:=200753849;
   	OWF_Key[306,7]:=1450403442;
   	OWF_Key[306,8]:=882557552;
   	OWF_Key[306,9]:=2025441160;
   	OWF_Key[306,10]:=2017827652;
   	OWF_Key[306,11]:=567324796;
   	OWF_Key[306,12]:=974302648;
   	OWF_Key[307,0]:=2092711674;
   	OWF_Key[307,1]:=2012740436;
   	OWF_Key[307,2]:=647780916;
   	OWF_Key[307,3]:=694158644;
   	OWF_Key[307,4]:=1431581549;
   	OWF_Key[307,5]:=1366437201;
   	OWF_Key[307,6]:=1386403931;
   	OWF_Key[307,7]:=40117105;
   	OWF_Key[307,8]:=1557715136;
   	OWF_Key[307,9]:=1389295347;
   	OWF_Key[307,10]:=585757347;
   	OWF_Key[307,11]:=849923725;
   	OWF_Key[307,12]:=1934760430;
   	OWF_Key[308,0]:=1722912930;
   	OWF_Key[308,1]:=989049945;
   	OWF_Key[308,2]:=1434792138;
   	OWF_Key[308,3]:=1795551986;
   	OWF_Key[308,4]:=545376040;
   	OWF_Key[308,5]:=932599939;
   	OWF_Key[308,6]:=403323632;
   	OWF_Key[308,7]:=1790466851;
   	OWF_Key[308,8]:=62625787;
   	OWF_Key[308,9]:=490336956;
   	OWF_Key[308,10]:=451154998;
   	OWF_Key[308,11]:=2015124611;
   	OWF_Key[308,12]:=1929430569;
   	OWF_Key[309,0]:=1373854605;
   	OWF_Key[309,1]:=1901562908;
   	OWF_Key[309,2]:=1305595762;
   	OWF_Key[309,3]:=1035847518;
   	OWF_Key[309,4]:=2077695225;
   	OWF_Key[309,5]:=1344844477;
   	OWF_Key[309,6]:=1010259473;
   	OWF_Key[309,7]:=922250580;
   	OWF_Key[309,8]:=1622875035;
   	OWF_Key[309,9]:=154427342;
   	OWF_Key[309,10]:=1175859706;
   	OWF_Key[309,11]:=94130927;
   	OWF_Key[309,12]:=1409996140;
   	OWF_Key[310,0]:=229565709;
   	OWF_Key[310,1]:=148723469;
   	OWF_Key[310,2]:=1727534663;
   	OWF_Key[310,3]:=1184917341;
   	OWF_Key[310,4]:=1071363996;
   	OWF_Key[310,5]:=443949111;
   	OWF_Key[310,6]:=506797285;
   	OWF_Key[310,7]:=1655431183;
   	OWF_Key[310,8]:=824685404;
   	OWF_Key[310,9]:=1600711337;
   	OWF_Key[310,10]:=587245000;
   	OWF_Key[310,11]:=1147194895;
   	OWF_Key[310,12]:=898888513;
   	OWF_Key[311,0]:=1854506430;
   	OWF_Key[311,1]:=438339574;
   	OWF_Key[311,2]:=1078153287;
   	OWF_Key[311,3]:=1499750094;
   	OWF_Key[311,4]:=1886362493;
   	OWF_Key[311,5]:=1805443847;
   	OWF_Key[311,6]:=1162745426;
   	OWF_Key[311,7]:=830263901;
   	OWF_Key[311,8]:=1063161141;
   	OWF_Key[311,9]:=620275595;
   	OWF_Key[311,10]:=1731504959;
   	OWF_Key[311,11]:=911334105;
   	OWF_Key[311,12]:=482497532;
   	OWF_Key[312,0]:=625162908;
   	OWF_Key[312,1]:=2102550000;
   	OWF_Key[312,2]:=405889591;
   	OWF_Key[312,3]:=332204328;
   	OWF_Key[312,4]:=1346018900;
   	OWF_Key[312,5]:=1836695371;
   	OWF_Key[312,6]:=1791877907;
   	OWF_Key[312,7]:=956132716;
   	OWF_Key[312,8]:=997749220;
   	OWF_Key[312,9]:=2015790650;
   	OWF_Key[312,10]:=2141741790;
   	OWF_Key[312,11]:=893721873;
   	OWF_Key[312,12]:=626685030;
   	OWF_Key[313,0]:=1922384603;
   	OWF_Key[313,1]:=1956752228;
   	OWF_Key[313,2]:=2029720698;
   	OWF_Key[313,3]:=1193903627;
   	OWF_Key[313,4]:=1760272519;
   	OWF_Key[313,5]:=668106909;
   	OWF_Key[313,6]:=1021138685;
   	OWF_Key[313,7]:=236982347;
   	OWF_Key[313,8]:=1576687950;